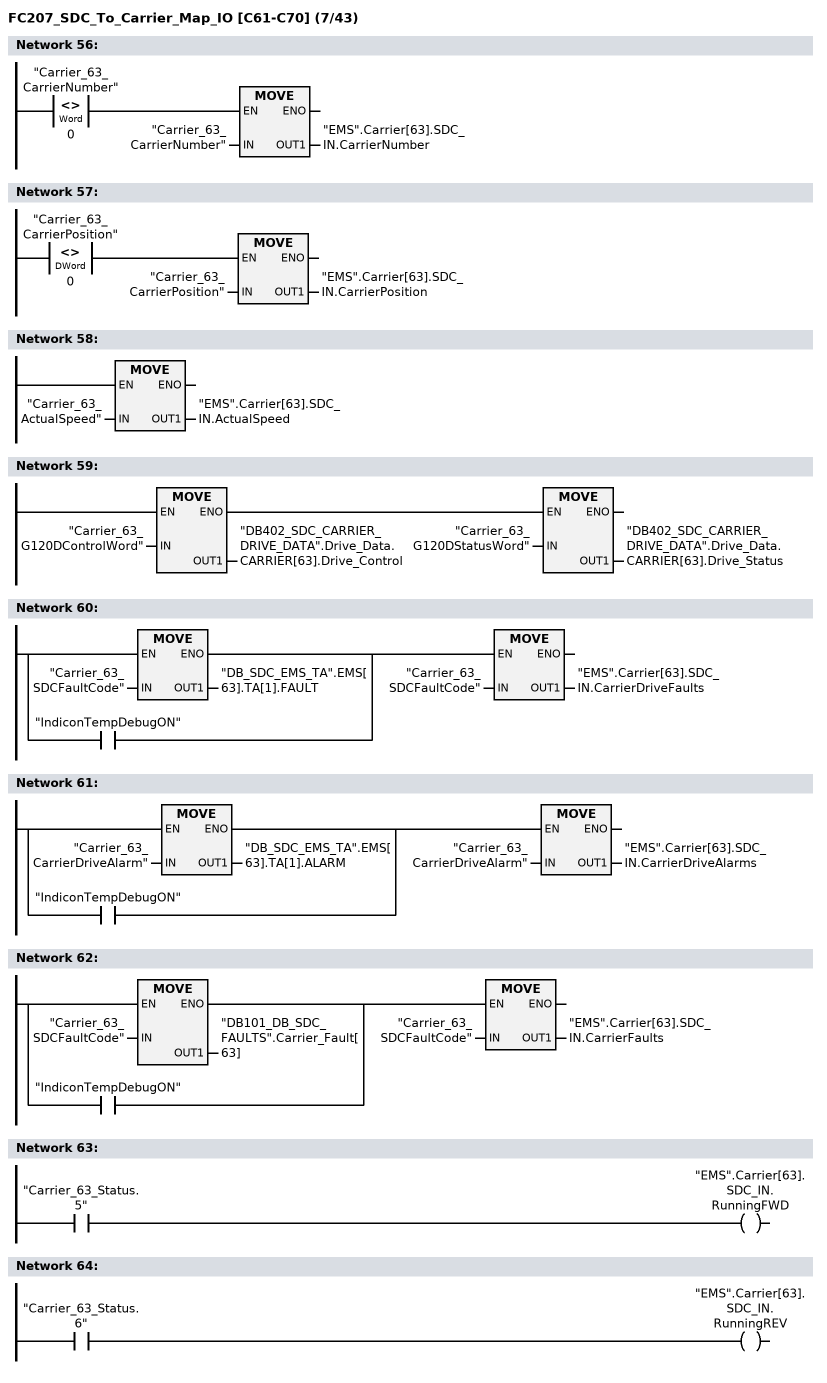
   RUNG wire#powerrail
      { S7_Templates := "SrcType := Word" } NE_Contact(in1 := "Carrier_63_CarrierNumber", in2 := 0)
      Move(in := "Carrier_63_CarrierNumber", out1 => "EMS".Carrier[63].SDC_IN.CarrierNumber)
   END_RUNG
   // the same network as SCL:
   IF "Carrier_63_CarrierNumber" <> 0 THEN
       "EMS".Carrier[63].SDC_IN.CarrierNumber := "Carrier_63_CarrierNumber";
   END_IF;
END_REGION

REGION Network 57
   RUNG wire#powerrail
      { S7_Templates := "SrcType := DWord" } NE_Contact(in1 := "Carrier_63_CarrierPosition", in2 := 0)
      Move(in := "Carrier_63_CarrierPosition", out1 => "EMS".Carrier[63].SDC_IN.CarrierPosition)
   END_RUNG
   // the same network as SCL:
   IF "Carrier_63_CarrierPosition" <> 0 THEN
       "EMS".Carrier[63].SDC_IN.CarrierPosition := "Carrier_63_CarrierPosition";
   END_IF;
END_REGION

REGION Network 58
   RUNG wire#powerrail
      Move(in := "Carrier_63_ActualSpeed", out1 => "EMS".Carrier[63].SDC_IN.ActualSpeed)
   END_RUNG
   // the same network as SCL:
   "EMS".Carrier[63].SDC_IN.ActualSpeed := "Carrier_63_ActualSpeed";
END_REGION

REGION Network 59
   RUNG wire#powerrail
      Move(in := "Carrier_63_G120DControlWord", out1 => "DB402_SDC_CARRIER_DRIVE_DATA".Drive_Data.CARRIER[63].Drive_Control)
      Move(in := "Carrier_63_G120DStatusWord", out1 => "DB402_SDC_CARRIER_DRIVE_DATA".Drive_Data.CARRIER[63].Drive_Status)
   END_RUNG
   // the same network as SCL:
   "DB402_SDC_CARRIER_DRIVE_DATA".Drive_Data.CARRIER[63].Drive_Control := "Carrier_63_G120DControlWord";
   "DB402_SDC_CARRIER_DRIVE_DATA".Drive_Data.CARRIER[63].Drive_Status := "Carrier_63_G120DStatusWord";
END_REGION

REGION Network 60
   RUNG wire#powerrail
      Move(in := "Carrier_63_SDCFaultCode", out1 => "DB_SDC_EMS_TA".EMS[63].TA[1].FAULT)
      wire#w1
      Move(in := "Carrier_63_SDCFaultCode", out1 => "EMS".Carrier[63].SDC_IN.CarrierDriveFaults)
   END_RUNG
   RUNG wire#powerrail
      Contact( "IndiconTempDebugON" )
   END_RUNG wire#w1
   // the same network as SCL:
   "DB_SDC_EMS_TA".EMS[63].TA[1].FAULT := "Carrier_63_SDCFaultCode";
   IF TRUE OR "IndiconTempDebugON" THEN
       "EMS".Carrier[63].SDC_IN.CarrierDriveFaults := "Carrier_63_SDCFaultCode";
   END_IF;
END_REGION

REGION Network 61
   RUNG wire#powerrail
      Move(in := "Carrier_63_CarrierDriveAlarm", out1 => "DB_SDC_EMS_TA".EMS[63].TA[1].ALARM)
      wire#w1
      Move(in := "Carrier_63_CarrierDriveAlarm", out1 => "EMS".Carrier[63].SDC_IN.CarrierDriveAlarms)
   END_RUNG
   RUNG wire#powerrail
      Contact( "IndiconTempDebugON" )
   END_RUNG wire#w1
   // the same network as SCL:
   "DB_SDC_EMS_TA".EMS[63].TA[1].ALARM := "Carrier_63_CarrierDriveAlarm";
   IF TRUE OR "IndiconTempDebugON" THEN
       "EMS".Carrier[63].SDC_IN.CarrierDriveAlarms := "Carrier_63_CarrierDriveAlarm";
   END_IF;
END_REGION

REGION Network 62
   RUNG wire#powerrail
      Move(in := "Carrier_63_SDCFaultCode", out1 => "DB101_DB_SDC_FAULTS".Carrier_Fault[63])
      wire#w1
      Move(in := "Carrier_63_SDCFaultCode", out1 => "EMS".Carrier[63].SDC_IN.CarrierFaults)
   END_RUNG
   RUNG wire#powerrail
      Contact( "IndiconTempDebugON" )
   END_RUNG wire#w1
   // the same network as SCL:
   "DB101_DB_SDC_FAULTS".Carrier_Fault[63] := "Carrier_63_SDCFaultCode";
   IF TRUE OR "IndiconTempDebugON" THEN
       "EMS".Carrier[63].SDC_IN.CarrierFaults := "Carrier_63_SDCFaultCode";
   END_IF;
END_REGION

REGION Network 63
   RUNG wire#powerrail
      Contact( "Carrier_63_Status.5" )
      Coil( "EMS".Carrier[63].SDC_IN.RunningFWD )
   END_RUNG
   // the same network as SCL:
   "EMS".Carrier[63].SDC_IN.RunningFWD := "Carrier_63_Status.5";
END_REGION

REGION Network 64
   RUNG wire#powerrail
      Contact( "Carrier_63_Status.6" )
      Coil( "EMS".Carrier[63].SDC_IN.RunningREV )
   END_RUNG
   // the same network as SCL:
   "EMS".Carrier[63].SDC_IN.RunningREV := "Carrier_63_Status.6";
END_REGION

REGION Network 65
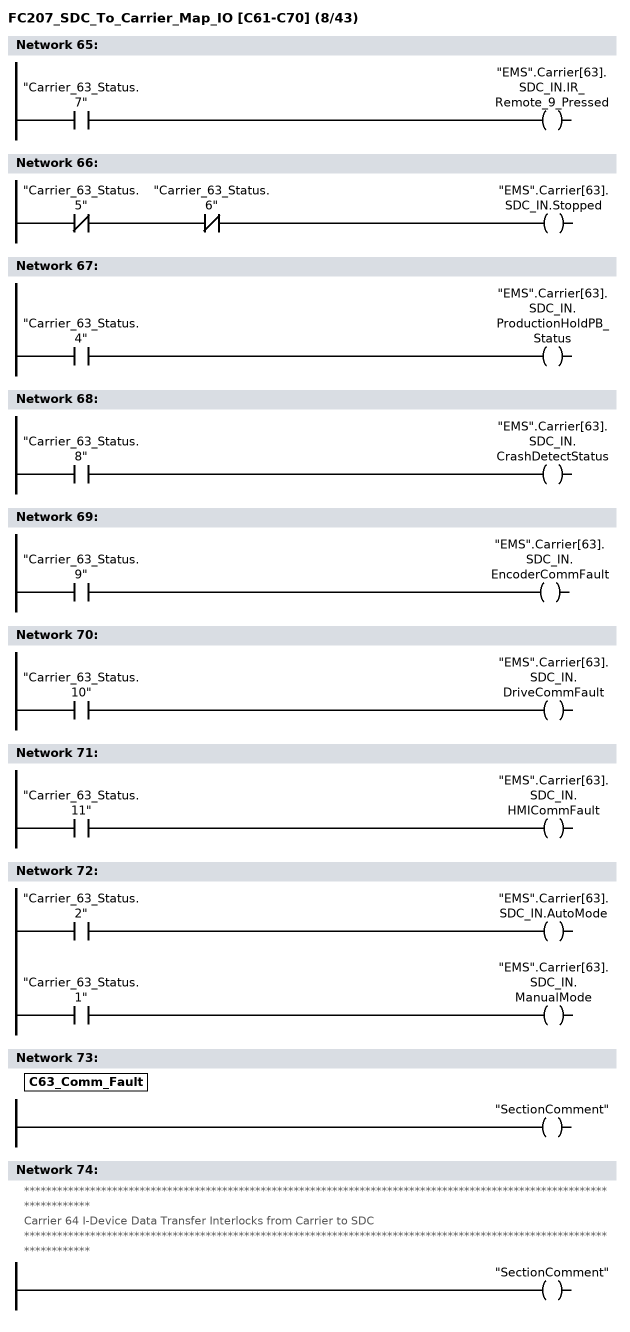
   RUNG wire#powerrail
      Contact( "Carrier_63_Status.7" )
      Coil( "EMS".Carrier[63].SDC_IN.IR_Remote_9_Pressed )
   END_RUNG
   // the same network as SCL:
   "EMS".Carrier[63].SDC_IN.IR_Remote_9_Pressed := "Carrier_63_Status.7";
END_REGION

REGION Network 66
   RUNG wire#powerrail
      I_Contact( "Carrier_63_Status.5" )
      I_Contact( "Carrier_63_Status.6" )
      Coil( "EMS".Carrier[63].SDC_IN.Stopped )
   END_RUNG
   // the same network as SCL:
   "EMS".Carrier[63].SDC_IN.Stopped := NOT "Carrier_63_Status.5" AND NOT "Carrier_63_Status.6";
END_REGION

REGION Network 67
   RUNG wire#powerrail
      Contact( "Carrier_63_Status.4" )
      Coil( "EMS".Carrier[63].SDC_IN.ProductionHoldPB_Status )
   END_RUNG
   // the same network as SCL:
   "EMS".Carrier[63].SDC_IN.ProductionHoldPB_Status := "Carrier_63_Status.4";
END_REGION

REGION Network 68
   RUNG wire#powerrail
      Contact( "Carrier_63_Status.8" )
      Coil( "EMS".Carrier[63].SDC_IN.CrashDetectStatus )
   END_RUNG
   // the same network as SCL:
   "EMS".Carrier[63].SDC_IN.CrashDetectStatus := "Carrier_63_Status.8";
END_REGION

REGION Network 69
   RUNG wire#powerrail
      Contact( "Carrier_63_Status.9" )
      Coil( "EMS".Carrier[63].SDC_IN.EncoderCommFault )
   END_RUNG
   // the same network as SCL:
   "EMS".Carrier[63].SDC_IN.EncoderCommFault := "Carrier_63_Status.9";
END_REGION

REGION Network 70
   RUNG wire#powerrail
      Contact( "Carrier_63_Status.10" )
      Coil( "EMS".Carrier[63].SDC_IN.DriveCommFault )
   END_RUNG
   // the same network as SCL:
   "EMS".Carrier[63].SDC_IN.DriveCommFault := "Carrier_63_Status.10";
END_REGION

REGION Network 71
   RUNG wire#powerrail
      Contact( "Carrier_63_Status.11" )
      Coil( "EMS".Carrier[63].SDC_IN.HMICommFault )
   END_RUNG
   // the same network as SCL:
   "EMS".Carrier[63].SDC_IN.HMICommFault := "Carrier_63_Status.11";
END_REGION

REGION Network 72
   RUNG wire#powerrail
      Contact( "Carrier_63_Status.2" )
      Coil( "EMS".Carrier[63].SDC_IN.AutoMode )
   END_RUNG
   RUNG wire#powerrail
      Contact( "Carrier_63_Status.1" )
      Coil( "EMS".Carrier[63].SDC_IN.ManualMode )
   END_RUNG
   // the same network as SCL:
   "EMS".Carrier[63].SDC_IN.AutoMode := "Carrier_63_Status.2";
   "EMS".Carrier[63].SDC_IN.ManualMode := "Carrier_63_Status.1";
END_REGION

REGION Network 73
   Label( C63_Comm_Fault )
   RUNG wire#powerrail
      Coil( "SectionComment" )
   END_RUNG
   // the same network as SCL:
   C63_Comm_Fault:
   "SectionComment" := TRUE;
END_REGION

REGION Network 74
   // **********************************************************************************************************************
   // 
   // Carrier 64 I-Device Data Transfer Interlocks from Carrier to SDC
   // 
   // **********************************************************************************************************************
   RUNG wire#powerrail
      Coil( "SectionComment" )
   END_RUNG
   // the same network as SCL:
   "SectionComment" := TRUE;
END_REGION

REGION Network 75
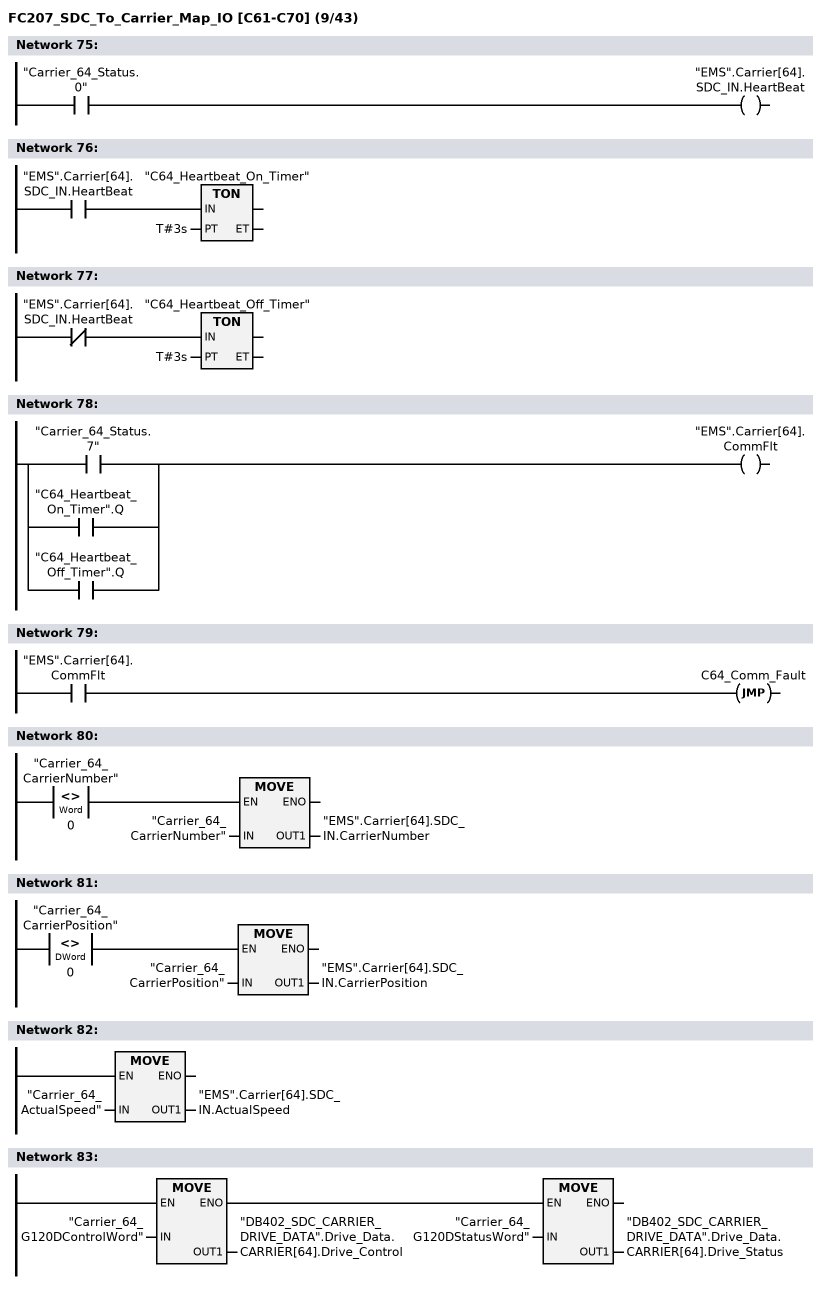
   RUNG wire#powerrail
      Contact( "Carrier_64_Status.0" )
      Coil( "EMS".Carrier[64].SDC_IN.HeartBeat )
   END_RUNG
   // the same network as SCL:
   "EMS".Carrier[64].SDC_IN.HeartBeat := "Carrier_64_Status.0";
END_REGION

REGION Network 76
   "C64_Heartbeat_On_Timer".TON(IN := "EMS".Carrier[64].SDC_IN.HeartBeat, PT := T#3s);
END_REGION

REGION Network 77
   "C64_Heartbeat_Off_Timer".TON(IN := NOT "EMS".Carrier[64].SDC_IN.HeartBeat, PT := T#3s);
END_REGION

REGION Network 78
   RUNG wire#powerrail
      Contact( "Carrier_64_Status.7" )
      wire#w1
      Coil( "EMS".Carrier[64].CommFlt )
   END_RUNG
   RUNG wire#powerrail
      Contact( "C64_Heartbeat_On_Timer".Q )
   END_RUNG wire#w1
   RUNG wire#powerrail
      Contact( "C64_Heartbeat_Off_Timer".Q )
   END_RUNG wire#w1
   // the same network as SCL:
   "EMS".Carrier[64].CommFlt := "Carrier_64_Status.7" OR "C64_Heartbeat_On_Timer".Q OR "C64_Heartbeat_Off_Timer".Q;
END_REGION

REGION Network 79
   RUNG wire#powerrail
      Contact( "EMS".Carrier[64].CommFlt )
      JumpCoil( C64_Comm_Fault )
   END_RUNG
   // the same network as SCL:
   IF "EMS".Carrier[64].CommFlt THEN GOTO C64_Comm_Fault; END_IF;
END_REGION

REGION Network 80
   RUNG wire#powerrail
      { S7_Templates := "SrcType := Word" } NE_Contact(in1 := "Carrier_64_CarrierNumber", in2 := 0)
      Move(in := "Carrier_64_CarrierNumber", out1 => "EMS".Carrier[64].SDC_IN.CarrierNumber)
   END_RUNG
   // the same network as SCL:
   IF "Carrier_64_CarrierNumber" <> 0 THEN
       "EMS".Carrier[64].SDC_IN.CarrierNumber := "Carrier_64_CarrierNumber";
   END_IF;
END_REGION

REGION Network 81
   RUNG wire#powerrail
      { S7_Templates := "SrcType := DWord" } NE_Contact(in1 := "Carrier_64_CarrierPosition", in2 := 0)
      Move(in := "Carrier_64_CarrierPosition", out1 => "EMS".Carrier[64].SDC_IN.CarrierPosition)
   END_RUNG
   // the same network as SCL:
   IF "Carrier_64_CarrierPosition" <> 0 THEN
       "EMS".Carrier[64].SDC_IN.CarrierPosition := "Carrier_64_CarrierPosition";
   END_IF;
END_REGION

REGION Network 82
   RUNG wire#powerrail
      Move(in := "Carrier_64_ActualSpeed", out1 => "EMS".Carrier[64].SDC_IN.ActualSpeed)
   END_RUNG
   // the same network as SCL:
   "EMS".Carrier[64].SDC_IN.ActualSpeed := "Carrier_64_ActualSpeed";
END_REGION

REGION Network 83
   RUNG wire#powerrail
      Move(in := "Carrier_64_G120DControlWord", out1 => "DB402_SDC_CARRIER_DRIVE_DATA".Drive_Data.CARRIER[64].Drive_Control)
      Move(in := "Carrier_64_G120DStatusWord", out1 => "DB402_SDC_CARRIER_DRIVE_DATA".Drive_Data.CARRIER[64].Drive_Status)
   END_RUNG
   // the same network as SCL:
   "DB402_SDC_CARRIER_DRIVE_DATA".Drive_Data.CARRIER[64].Drive_Control := "Carrier_64_G120DControlWord";
   "DB402_SDC_CARRIER_DRIVE_DATA".Drive_Data.CARRIER[64].Drive_Status := "Carrier_64_G120DStatusWord";
END_REGION

REGION Network 84
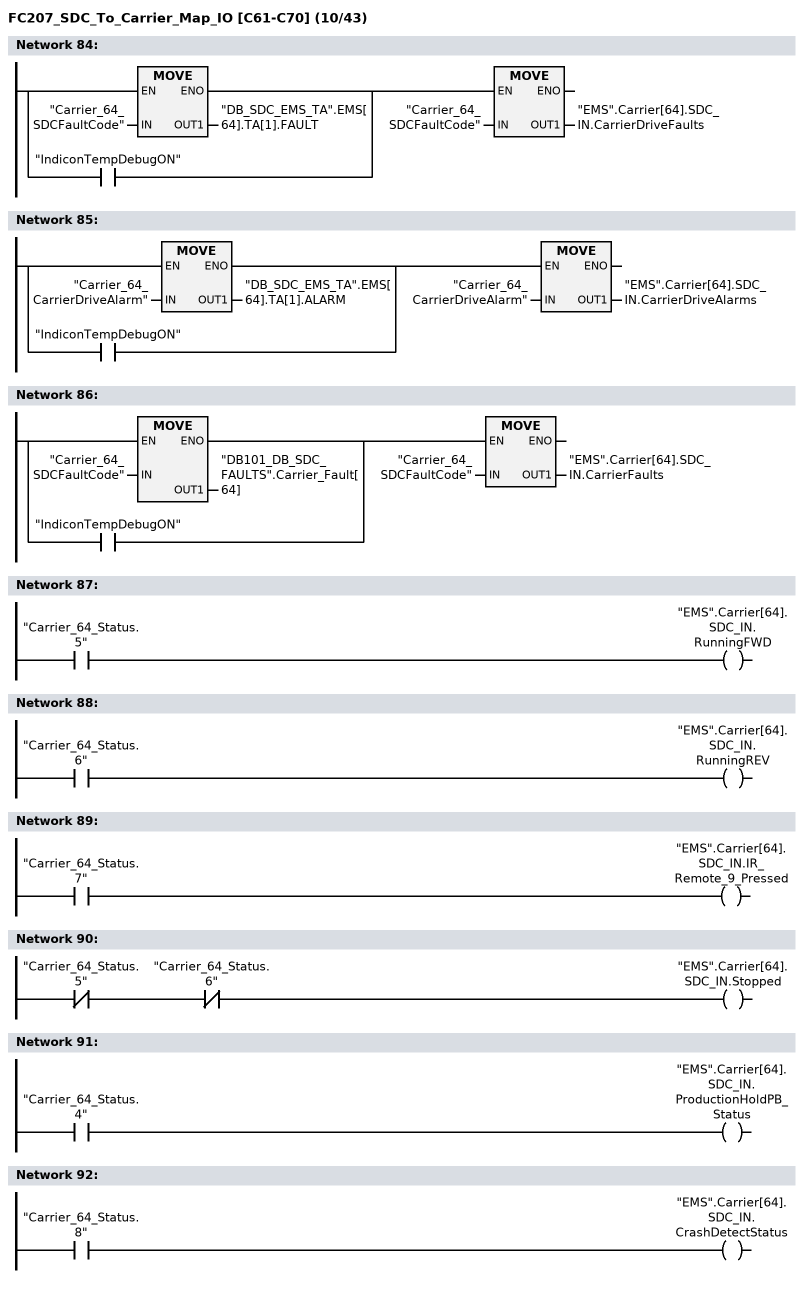
   RUNG wire#powerrail
      Move(in := "Carrier_64_SDCFaultCode", out1 => "DB_SDC_EMS_TA".EMS[64].TA[1].FAULT)
      wire#w1
      Move(in := "Carrier_64_SDCFaultCode", out1 => "EMS".Carrier[64].SDC_IN.CarrierDriveFaults)
   END_RUNG
   RUNG wire#powerrail
      Contact( "IndiconTempDebugON" )
   END_RUNG wire#w1
   // the same network as SCL:
   "DB_SDC_EMS_TA".EMS[64].TA[1].FAULT := "Carrier_64_SDCFaultCode";
   IF TRUE OR "IndiconTempDebugON" THEN
       "EMS".Carrier[64].SDC_IN.CarrierDriveFaults := "Carrier_64_SDCFaultCode";
   END_IF;
END_REGION

REGION Network 85
   RUNG wire#powerrail
      Move(in := "Carrier_64_CarrierDriveAlarm", out1 => "DB_SDC_EMS_TA".EMS[64].TA[1].ALARM)
      wire#w1
      Move(in := "Carrier_64_CarrierDriveAlarm", out1 => "EMS".Carrier[64].SDC_IN.CarrierDriveAlarms)
   END_RUNG
   RUNG wire#powerrail
      Contact( "IndiconTempDebugON" )
   END_RUNG wire#w1
   // the same network as SCL:
   "DB_SDC_EMS_TA".EMS[64].TA[1].ALARM := "Carrier_64_CarrierDriveAlarm";
   IF TRUE OR "IndiconTempDebugON" THEN
       "EMS".Carrier[64].SDC_IN.CarrierDriveAlarms := "Carrier_64_CarrierDriveAlarm";
   END_IF;
END_REGION

REGION Network 86
   RUNG wire#powerrail
      Move(in := "Carrier_64_SDCFaultCode", out1 => "DB101_DB_SDC_FAULTS".Carrier_Fault[64])
      wire#w1
      Move(in := "Carrier_64_SDCFaultCode", out1 => "EMS".Carrier[64].SDC_IN.CarrierFaults)
   END_RUNG
   RUNG wire#powerrail
      Contact( "IndiconTempDebugON" )
   END_RUNG wire#w1
   // the same network as SCL:
   "DB101_DB_SDC_FAULTS".Carrier_Fault[64] := "Carrier_64_SDCFaultCode";
   IF TRUE OR "IndiconTempDebugON" THEN
       "EMS".Carrier[64].SDC_IN.CarrierFaults := "Carrier_64_SDCFaultCode";
   END_IF;
END_REGION

REGION Network 87
   RUNG wire#powerrail
      Contact( "Carrier_64_Status.5" )
      Coil( "EMS".Carrier[64].SDC_IN.RunningFWD )
   END_RUNG
   // the same network as SCL:
   "EMS".Carrier[64].SDC_IN.RunningFWD := "Carrier_64_Status.5";
END_REGION

REGION Network 88
   RUNG wire#powerrail
      Contact( "Carrier_64_Status.6" )
      Coil( "EMS".Carrier[64].SDC_IN.RunningREV )
   END_RUNG
   // the same network as SCL:
   "EMS".Carrier[64].SDC_IN.RunningREV := "Carrier_64_Status.6";
END_REGION

REGION Network 89
   RUNG wire#powerrail
      Contact( "Carrier_64_Status.7" )
      Coil( "EMS".Carrier[64].SDC_IN.IR_Remote_9_Pressed )
   END_RUNG
   // the same network as SCL:
   "EMS".Carrier[64].SDC_IN.IR_Remote_9_Pressed := "Carrier_64_Status.7";
END_REGION

REGION Network 90
   RUNG wire#powerrail
      I_Contact( "Carrier_64_Status.5" )
      I_Contact( "Carrier_64_Status.6" )
      Coil( "EMS".Carrier[64].SDC_IN.Stopped )
   END_RUNG
   // the same network as SCL:
   "EMS".Carrier[64].SDC_IN.Stopped := NOT "Carrier_64_Status.5" AND NOT "Carrier_64_Status.6";
END_REGION

REGION Network 91
   RUNG wire#powerrail
      Contact( "Carrier_64_Status.4" )
      Coil( "EMS".Carrier[64].SDC_IN.ProductionHoldPB_Status )
   END_RUNG
   // the same network as SCL:
   "EMS".Carrier[64].SDC_IN.ProductionHoldPB_Status := "Carrier_64_Status.4";
END_REGION

REGION Network 92
   RUNG wire#powerrail
      Contact( "Carrier_64_Status.8" )
      Coil( "EMS".Carrier[64].SDC_IN.CrashDetectStatus )
   END_RUNG
   // the same network as SCL:
   "EMS".Carrier[64].SDC_IN.CrashDetectStatus := "Carrier_64_Status.8";
END_REGION

REGION Network 93
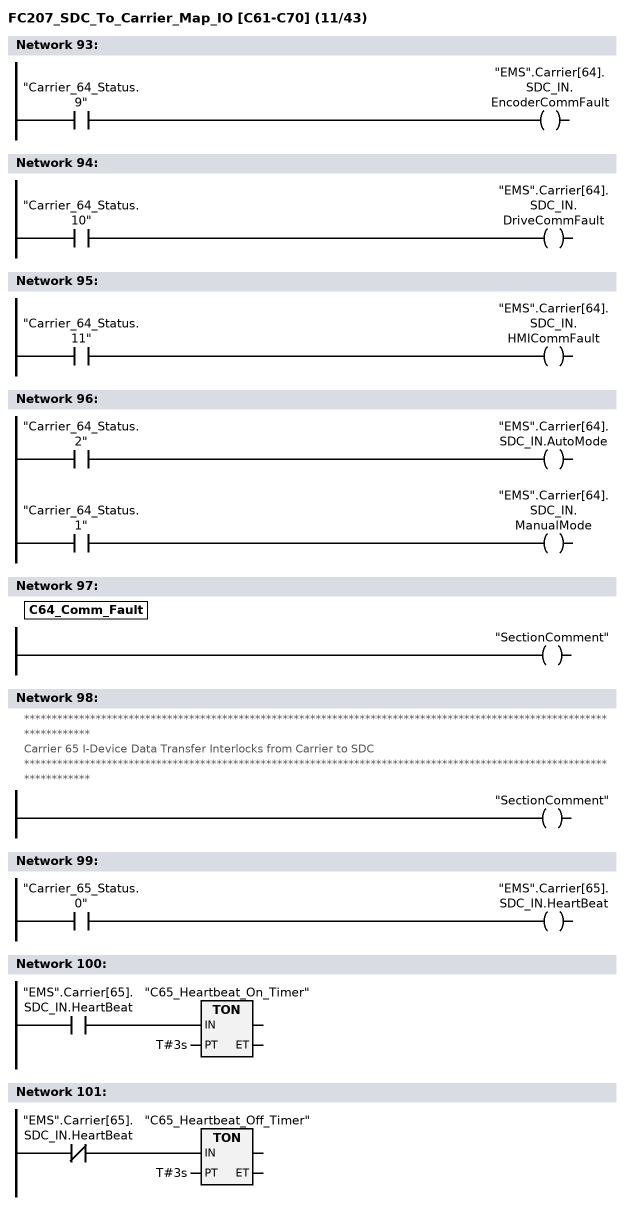
   RUNG wire#powerrail
      Contact( "Carrier_64_Status.9" )
      Coil( "EMS".Carrier[64].SDC_IN.EncoderCommFault )
   END_RUNG
   // the same network as SCL:
   "EMS".Carrier[64].SDC_IN.EncoderCommFault := "Carrier_64_Status.9";
END_REGION

REGION Network 94
   RUNG wire#powerrail
      Contact( "Carrier_64_Status.10" )
      Coil( "EMS".Carrier[64].SDC_IN.DriveCommFault )
   END_RUNG
   // the same network as SCL:
   "EMS".Carrier[64].SDC_IN.DriveCommFault := "Carrier_64_Status.10";
END_REGION

REGION Network 95
   RUNG wire#powerrail
      Contact( "Carrier_64_Status.11" )
      Coil( "EMS".Carrier[64].SDC_IN.HMICommFault )
   END_RUNG
   // the same network as SCL:
   "EMS".Carrier[64].SDC_IN.HMICommFault := "Carrier_64_Status.11";
END_REGION

REGION Network 96
   RUNG wire#powerrail
      Contact( "Carrier_64_Status.2" )
      Coil( "EMS".Carrier[64].SDC_IN.AutoMode )
   END_RUNG
   RUNG wire#powerrail
      Contact( "Carrier_64_Status.1" )
      Coil( "EMS".Carrier[64].SDC_IN.ManualMode )
   END_RUNG
   // the same network as SCL:
   "EMS".Carrier[64].SDC_IN.AutoMode := "Carrier_64_Status.2";
   "EMS".Carrier[64].SDC_IN.ManualMode := "Carrier_64_Status.1";
END_REGION

REGION Network 97
   Label( C64_Comm_Fault )
   RUNG wire#powerrail
      Coil( "SectionComment" )
   END_RUNG
   // the same network as SCL:
   C64_Comm_Fault:
   "SectionComment" := TRUE;
END_REGION

REGION Network 98
   // **********************************************************************************************************************
   // 
   // Carrier 65 I-Device Data Transfer Interlocks from Carrier to SDC
   // 
   // **********************************************************************************************************************
   RUNG wire#powerrail
      Coil( "SectionComment" )
   END_RUNG
   // the same network as SCL:
   "SectionComment" := TRUE;
END_REGION

REGION Network 99
   RUNG wire#powerrail
      Contact( "Carrier_65_Status.0" )
      Coil( "EMS".Carrier[65].SDC_IN.HeartBeat )
   END_RUNG
   // the same network as SCL:
   "EMS".Carrier[65].SDC_IN.HeartBeat := "Carrier_65_Status.0";
END_REGION

REGION Network 100
   "C65_Heartbeat_On_Timer".TON(IN := "EMS".Carrier[65].SDC_IN.HeartBeat, PT := T#3s);
END_REGION

REGION Network 101
   "C65_Heartbeat_Off_Timer".TON(IN := NOT "EMS".Carrier[65].SDC_IN.HeartBeat, PT := T#3s);
END_REGION

REGION Network 102
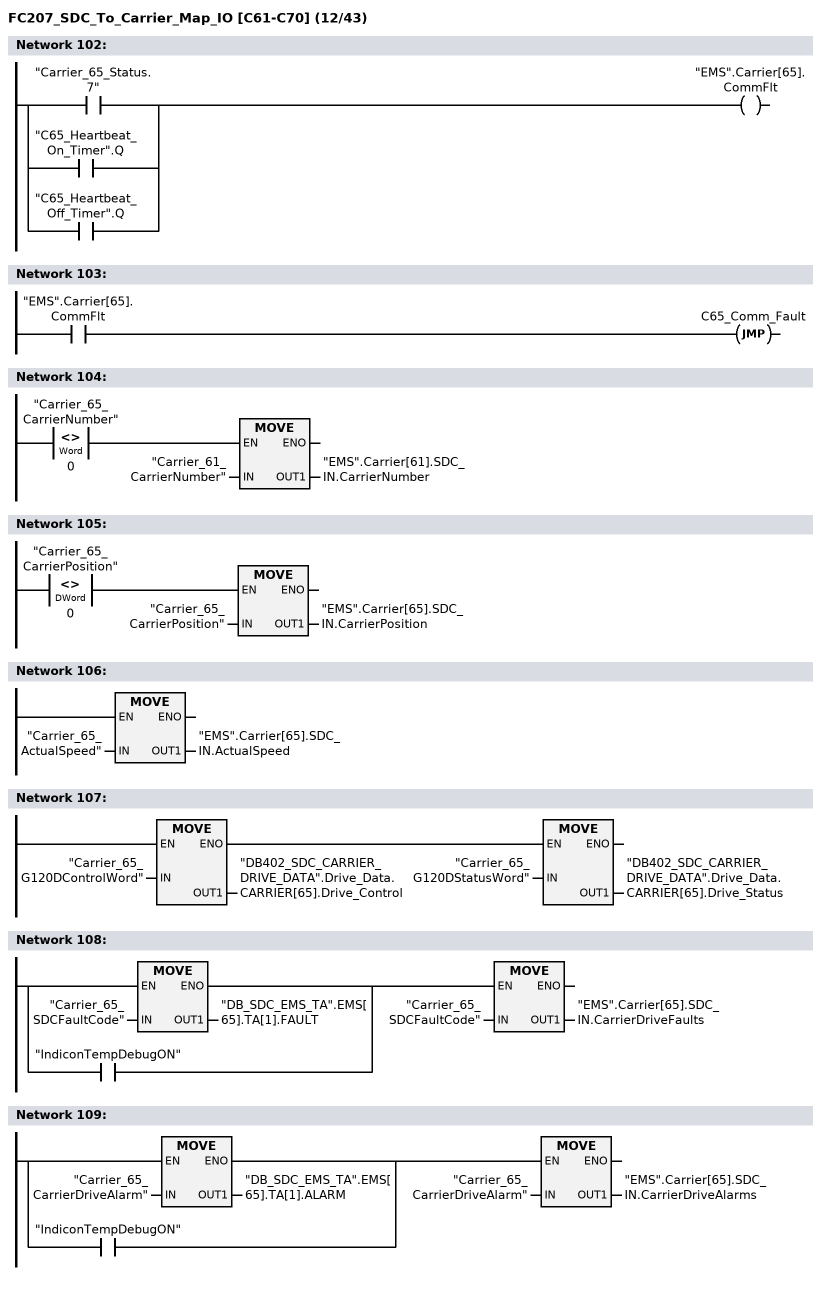
   RUNG wire#powerrail
      Contact( "Carrier_65_Status.7" )
      wire#w1
      Coil( "EMS".Carrier[65].CommFlt )
   END_RUNG
   RUNG wire#powerrail
      Contact( "C65_Heartbeat_On_Timer".Q )
   END_RUNG wire#w1
   RUNG wire#powerrail
      Contact( "C65_Heartbeat_Off_Timer".Q )
   END_RUNG wire#w1
   // the same network as SCL:
   "EMS".Carrier[65].CommFlt := "Carrier_65_Status.7" OR "C65_Heartbeat_On_Timer".Q OR "C65_Heartbeat_Off_Timer".Q;
END_REGION

REGION Network 103
   RUNG wire#powerrail
      Contact( "EMS".Carrier[65].CommFlt )
      JumpCoil( C65_Comm_Fault )
   END_RUNG
   // the same network as SCL:
   IF "EMS".Carrier[65].CommFlt THEN GOTO C65_Comm_Fault; END_IF;
END_REGION

REGION Network 104
   RUNG wire#powerrail
      { S7_Templates := "SrcType := Word" } NE_Contact(in1 := "Carrier_65_CarrierNumber", in2 := 0)
      Move(in := "Carrier_61_CarrierNumber", out1 => "EMS".Carrier[61].SDC_IN.CarrierNumber)
   END_RUNG
   // the same network as SCL:
   IF "Carrier_65_CarrierNumber" <> 0 THEN
       "EMS".Carrier[61].SDC_IN.CarrierNumber := "Carrier_61_CarrierNumber";
   END_IF;
END_REGION

REGION Network 105
   RUNG wire#powerrail
      { S7_Templates := "SrcType := DWord" } NE_Contact(in1 := "Carrier_65_CarrierPosition", in2 := 0)
      Move(in := "Carrier_65_CarrierPosition", out1 => "EMS".Carrier[65].SDC_IN.CarrierPosition)
   END_RUNG
   // the same network as SCL:
   IF "Carrier_65_CarrierPosition" <> 0 THEN
       "EMS".Carrier[65].SDC_IN.CarrierPosition := "Carrier_65_CarrierPosition";
   END_IF;
END_REGION

REGION Network 106
   RUNG wire#powerrail
      Move(in := "Carrier_65_ActualSpeed", out1 => "EMS".Carrier[65].SDC_IN.ActualSpeed)
   END_RUNG
   // the same network as SCL:
   "EMS".Carrier[65].SDC_IN.ActualSpeed := "Carrier_65_ActualSpeed";
END_REGION

REGION Network 107
   RUNG wire#powerrail
      Move(in := "Carrier_65_G120DControlWord", out1 => "DB402_SDC_CARRIER_DRIVE_DATA".Drive_Data.CARRIER[65].Drive_Control)
      Move(in := "Carrier_65_G120DStatusWord", out1 => "DB402_SDC_CARRIER_DRIVE_DATA".Drive_Data.CARRIER[65].Drive_Status)
   END_RUNG
   // the same network as SCL:
   "DB402_SDC_CARRIER_DRIVE_DATA".Drive_Data.CARRIER[65].Drive_Control := "Carrier_65_G120DControlWord";
   "DB402_SDC_CARRIER_DRIVE_DATA".Drive_Data.CARRIER[65].Drive_Status := "Carrier_65_G120DStatusWord";
END_REGION

REGION Network 108
   RUNG wire#powerrail
      Move(in := "Carrier_65_SDCFaultCode", out1 => "DB_SDC_EMS_TA".EMS[65].TA[1].FAULT)
      wire#w1
      Move(in := "Carrier_65_SDCFaultCode", out1 => "EMS".Carrier[65].SDC_IN.CarrierDriveFaults)
   END_RUNG
   RUNG wire#powerrail
      Contact( "IndiconTempDebugON" )
   END_RUNG wire#w1
   // the same network as SCL:
   "DB_SDC_EMS_TA".EMS[65].TA[1].FAULT := "Carrier_65_SDCFaultCode";
   IF TRUE OR "IndiconTempDebugON" THEN
       "EMS".Carrier[65].SDC_IN.CarrierDriveFaults := "Carrier_65_SDCFaultCode";
   END_IF;
END_REGION

REGION Network 109
   RUNG wire#powerrail
      Move(in := "Carrier_65_CarrierDriveAlarm", out1 => "DB_SDC_EMS_TA".EMS[65].TA[1].ALARM)
      wire#w1
      Move(in := "Carrier_65_CarrierDriveAlarm", out1 => "EMS".Carrier[65].SDC_IN.CarrierDriveAlarms)
   END_RUNG
   RUNG wire#powerrail
      Contact( "IndiconTempDebugON" )
   END_RUNG wire#w1
   // the same network as SCL:
   "DB_SDC_EMS_TA".EMS[65].TA[1].ALARM := "Carrier_65_CarrierDriveAlarm";
   IF TRUE OR "IndiconTempDebugON" THEN
       "EMS".Carrier[65].SDC_IN.CarrierDriveAlarms := "Carrier_65_CarrierDriveAlarm";
   END_IF;
END_REGION

REGION Network 110
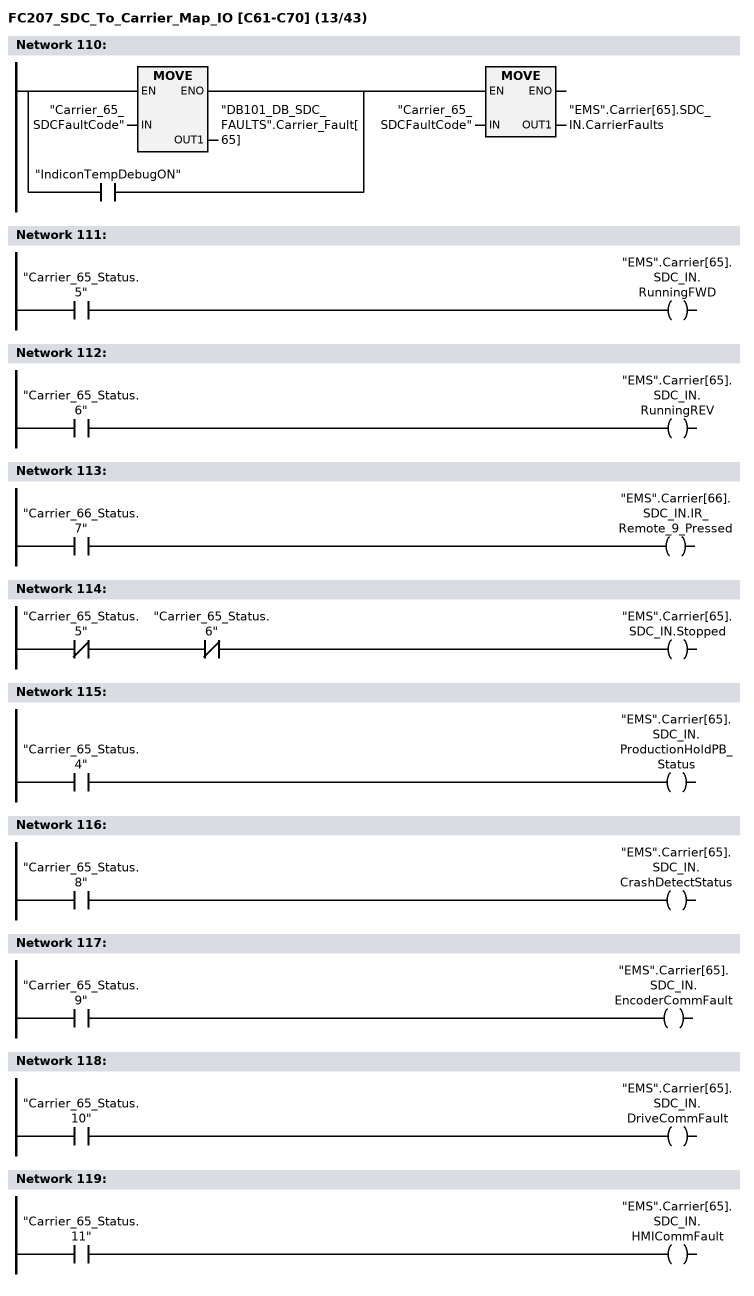
   RUNG wire#powerrail
      Move(in := "Carrier_65_SDCFaultCode", out1 => "DB101_DB_SDC_FAULTS".Carrier_Fault[65])
      wire#w1
      Move(in := "Carrier_65_SDCFaultCode", out1 => "EMS".Carrier[65].SDC_IN.CarrierFaults)
   END_RUNG
   RUNG wire#powerrail
      Contact( "IndiconTempDebugON" )
   END_RUNG wire#w1
   // the same network as SCL:
   "DB101_DB_SDC_FAULTS".Carrier_Fault[65] := "Carrier_65_SDCFaultCode";
   IF TRUE OR "IndiconTempDebugON" THEN
       "EMS".Carrier[65].SDC_IN.CarrierFaults := "Carrier_65_SDCFaultCode";
   END_IF;
END_REGION

REGION Network 111
   RUNG wire#powerrail
      Contact( "Carrier_65_Status.5" )
      Coil( "EMS".Carrier[65].SDC_IN.RunningFWD )
   END_RUNG
   // the same network as SCL:
   "EMS".Carrier[65].SDC_IN.RunningFWD := "Carrier_65_Status.5";
END_REGION

REGION Network 112
   RUNG wire#powerrail
      Contact( "Carrier_65_Status.6" )
      Coil( "EMS".Carrier[65].SDC_IN.RunningREV )
   END_RUNG
   // the same network as SCL:
   "EMS".Carrier[65].SDC_IN.RunningREV := "Carrier_65_Status.6";
END_REGION

REGION Network 113
   RUNG wire#powerrail
      Contact( "Carrier_66_Status.7" )
      Coil( "EMS".Carrier[66].SDC_IN.IR_Remote_9_Pressed )
   END_RUNG
   // the same network as SCL:
   "EMS".Carrier[66].SDC_IN.IR_Remote_9_Pressed := "Carrier_66_Status.7";
END_REGION

REGION Network 114
   RUNG wire#powerrail
      I_Contact( "Carrier_65_Status.5" )
      I_Contact( "Carrier_65_Status.6" )
      Coil( "EMS".Carrier[65].SDC_IN.Stopped )
   END_RUNG
   // the same network as SCL:
   "EMS".Carrier[65].SDC_IN.Stopped := NOT "Carrier_65_Status.5" AND NOT "Carrier_65_Status.6";
END_REGION

REGION Network 115
   RUNG wire#powerrail
      Contact( "Carrier_65_Status.4" )
      Coil( "EMS".Carrier[65].SDC_IN.ProductionHoldPB_Status )
   END_RUNG
   // the same network as SCL:
   "EMS".Carrier[65].SDC_IN.ProductionHoldPB_Status := "Carrier_65_Status.4";
END_REGION

REGION Network 116
   RUNG wire#powerrail
      Contact( "Carrier_65_Status.8" )
      Coil( "EMS".Carrier[65].SDC_IN.CrashDetectStatus )
   END_RUNG
   // the same network as SCL:
   "EMS".Carrier[65].SDC_IN.CrashDetectStatus := "Carrier_65_Status.8";
END_REGION

REGION Network 117
   RUNG wire#powerrail
      Contact( "Carrier_65_Status.9" )
      Coil( "EMS".Carrier[65].SDC_IN.EncoderCommFault )
   END_RUNG
   // the same network as SCL:
   "EMS".Carrier[65].SDC_IN.EncoderCommFault := "Carrier_65_Status.9";
END_REGION

REGION Network 118
   RUNG wire#powerrail
      Contact( "Carrier_65_Status.10" )
      Coil( "EMS".Carrier[65].SDC_IN.DriveCommFault )
   END_RUNG
   // the same network as SCL:
   "EMS".Carrier[65].SDC_IN.DriveCommFault := "Carrier_65_Status.10";
END_REGION

REGION Network 119
   RUNG wire#powerrail
      Contact( "Carrier_65_Status.11" )
      Coil( "EMS".Carrier[65].SDC_IN.HMICommFault )
   END_RUNG
   // the same network as SCL:
   "EMS".Carrier[65].SDC_IN.HMICommFault := "Carrier_65_Status.11";
END_REGION

REGION Network 120
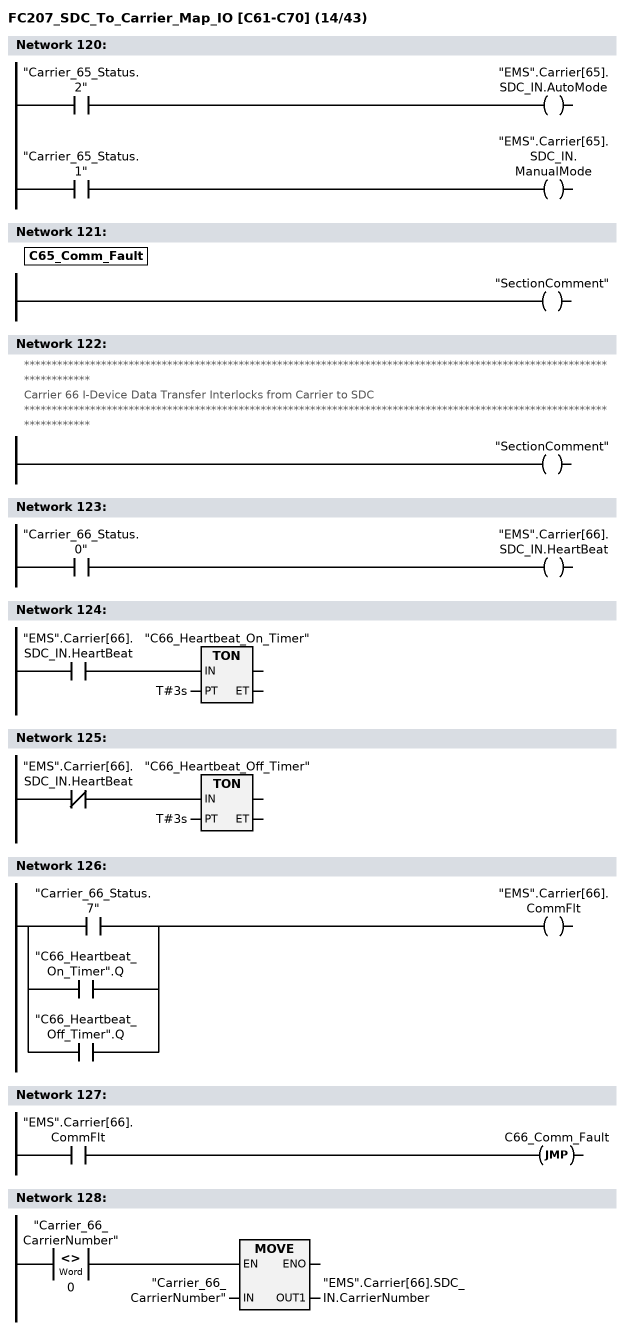
   RUNG wire#powerrail
      Contact( "Carrier_65_Status.2" )
      Coil( "EMS".Carrier[65].SDC_IN.AutoMode )
   END_RUNG
   RUNG wire#powerrail
      Contact( "Carrier_65_Status.1" )
      Coil( "EMS".Carrier[65].SDC_IN.ManualMode )
   END_RUNG
   // the same network as SCL:
   "EMS".Carrier[65].SDC_IN.AutoMode := "Carrier_65_Status.2";
   "EMS".Carrier[65].SDC_IN.ManualMode := "Carrier_65_Status.1";
END_REGION

REGION Network 121
   Label( C65_Comm_Fault )
   RUNG wire#powerrail
      Coil( "SectionComment" )
   END_RUNG
   // the same network as SCL:
   C65_Comm_Fault:
   "SectionComment" := TRUE;
END_REGION

REGION Network 122
   // **********************************************************************************************************************
   // 
   // Carrier 66 I-Device Data Transfer Interlocks from Carrier to SDC
   // 
   // **********************************************************************************************************************
   RUNG wire#powerrail
      Coil( "SectionComment" )
   END_RUNG
   // the same network as SCL:
   "SectionComment" := TRUE;
END_REGION

REGION Network 123
   RUNG wire#powerrail
      Contact( "Carrier_66_Status.0" )
      Coil( "EMS".Carrier[66].SDC_IN.HeartBeat )
   END_RUNG
   // the same network as SCL:
   "EMS".Carrier[66].SDC_IN.HeartBeat := "Carrier_66_Status.0";
END_REGION

REGION Network 124
   "C66_Heartbeat_On_Timer".TON(IN := "EMS".Carrier[66].SDC_IN.HeartBeat, PT := T#3s);
END_REGION

REGION Network 125
   "C66_Heartbeat_Off_Timer".TON(IN := NOT "EMS".Carrier[66].SDC_IN.HeartBeat, PT := T#3s);
END_REGION

REGION Network 126
   RUNG wire#powerrail
      Contact( "Carrier_66_Status.7" )
      wire#w1
      Coil( "EMS".Carrier[66].CommFlt )
   END_RUNG
   RUNG wire#powerrail
      Contact( "C66_Heartbeat_On_Timer".Q )
   END_RUNG wire#w1
   RUNG wire#powerrail
      Contact( "C66_Heartbeat_Off_Timer".Q )
   END_RUNG wire#w1
   // the same network as SCL:
   "EMS".Carrier[66].CommFlt := "Carrier_66_Status.7" OR "C66_Heartbeat_On_Timer".Q OR "C66_Heartbeat_Off_Timer".Q;
END_REGION

REGION Network 127
   RUNG wire#powerrail
      Contact( "EMS".Carrier[66].CommFlt )
      JumpCoil( C66_Comm_Fault )
   END_RUNG
   // the same network as SCL:
   IF "EMS".Carrier[66].CommFlt THEN GOTO C66_Comm_Fault; END_IF;
END_REGION
